// TIA Portal project "Lagerregal_1" (V20)

(* hardware
DEVICE "S7-1500/ET200MP-Station_1"  S7-1500 station
   slot 0: "Profilschiene_0"  Rack  6ES7 590-1***0-0AA0
   slot 1: "PLC_1"  CPU 1513-1 PN  6ES7 513-1AM03-0AB0  V4.0
      slot 3: "CPU-Display_1"  6ES7591-1AA00-0AA0
      slot 32768: "PROFINET-Schnittstelle_1"  X1
         slot 32769: "Port_1"  X1 P1
         slot 32770: "Port_2"  X1 P2
      slot 34817: "Virtual CP interface port_1"  Virtual CP interface port  Virtual CP interface port FW V4.0
   slot 2: "DI 16x24VDC BA_1"  DI 16x24VDC BA  6ES7 521-1BH10-0AA0  V1.1
   slot 3: "DQ 16x24VDC/0.5A ST_1"  DQ 16x24VDC/0.5A ST  6ES7 522-1BH00-0AB0  V2.0
   slot 4: "AI 8xU/I/R/RTD BA_2"  AI 8xU/I/R/RTD BA  6ES7 531-7QF00-0AB0  V1.0
   slot 5: "AI 8xU/I/R/RTD BA_1"  AI 8xU/I/R/RTD BA  6ES7 531-7QF00-0AB0  V1.0
DEVICE "HMI_1"  TP700 Comfort
   slot 0: "HMI_1"  TP700 Comfort  6AV2 124-0GC01-0AX0  17.0.0.0
   slot 1: "HMI_RT_1"  TP700 Comfort  6AV2 124-0GC01-0AX0  17.0.0.0
   slot 5: "HMI_1.IE_CP_1"  PROFINET Interface  17.0.0.0
      slot 1: "PROFINET Schnittstelle_1"  PROFINET Interface
         slot 1: "Port_1"  Port
         slot 2: "Port_2"  Port
   slot 7: "HMI_1.MPI/DP_CP_1"  MPI/DP Interface  17.0.0.0
*)

// ===== PLC "PLC_1"  CPU 1513-1 PN =====

VAR_GLOBAL   // PLC tag table "Variablentabelle aus XML_1"
   "E0.0 Not-Aus (S1)" AT %I0.0 : Bool;
   "E0.1 Anlage ein (S2)" AT %I0.1 : Bool;
   "E0.2 Start (S3)" AT %I0.2 : Bool;
   "E0.3 Sensor_Ein_SS (1B1)" AT %I0.3 : Bool;
   "E0.4 Sensor_Ein_SE (1B2)" AT %I0.4 : Bool;
   "E0.5 Sensor_Ein_MS (2B1)" AT %I0.5 : Bool;
   "E0.6 Sensor_Ein_ME (2B2)" AT %I0.6 : Bool;
   "E0.7 Sensor_Ein_EE (3B1)" AT %I0.7 : Bool;
   "E1.0 Sensor_Aus_S (4B1)" AT %I1.0 : Bool;
   "E1.1 Sensor_Aus_A (5B1)" AT %I1.1 : Bool;
   "E1.2 Kran_Gabel_Endlage (links) (6B1)" AT %I1.2 : Bool;
   "E1.3 Kran_Gabel_Endlage (rechts) (6B2)" AT %I1.3 : Bool;
   "E1.4 Kran_Gabel_Endage (mitte) (6B3)" AT %I1.4 : Bool;
   "E1.5 Kran_Gabel_Endlage (links) (7B1)" AT %I1.5 : Bool;
   "E1.6 Kran_Gabel_Endlage (rechts) (7B2)" AT %I1.6 : Bool;
   "E1.7 Kran_Gabel_Endage (mitte) (7B3)" AT %I1.7 : Bool;
   "A0.2 Start (H3)" AT %Q0.2 : Bool;
   "A0.3 Band_Ein_1 (1M1)" AT %Q0.3 : Bool;
   "A0.5 Band_Ein_2 (2M1)" AT %Q0.5 : Bool;
   "A0.7 Band_Ein_3 (3M1)" AT %Q0.7 : Bool;
   "A1.0 Band_Aus_1 (4M1)" AT %Q1.0 : Bool;
   "A1.1 Band_Aus_2 (5M1)" AT %Q1.1 : Bool;
   "A1.2 Kran_Gabel (links) (6M1)" AT %Q1.2 : Bool;
   "A1.3 Kran_Gabel (rechts) (6M2)" AT %Q1.3 : Bool;
   "A1.5 Kran_Gabel (links) (7M1)" AT %Q1.5 : Bool;
   "A1.6 Kran_Gabel (rechts) (7M2)" AT %Q1.6 : Bool;
   "EW30 Kamera (2B1)" AT %EW30 : Int;
   "EW34 Kran_Ist-X-Pos (6B4)" AT %EW32 : Int;
   "EW38 Kran_Ist-Z-Pos (6B5)" AT %EW34 : Int;
   "EW42 Kran_Ist-X-Pos (7B4)" AT %EW36 : Int;
   "EW46 Kran_Ist-Z-Pos (7B5)" AT %EW38 : Int;
   "AW34 Kran_Soll-X-Pos (6M4)" AT %AW32 : Int;
   "AW38 Kran_Soll-Z-Pos (6M5)" AT %AW34 : Int;
   "AW42 Kran_Soll-X-Pos (7M4)" AT %AW36 : Int;
   "AW46 Kran_Soll-Z-Pos (7M5)" AT %AW38 : Int;
END_VAR

TYPE "typKran_Pos"
   STRUCT
      "X-Ist" : Int;
      "X-Soll" : Int;
      "Z-Ist" : Int;
      "Z-Soll" : Int;
   END_STRUCT;
END_TYPE

TYPE "typLagerplatz"
   STRUCT
      Pos : Struct
         X : Int;
         Z : Int;
      END_STRUCT;
      Flags : Struct
         Belegt : Bool;
         In_Benutzung : Bool;
      END_STRUCT;
   END_STRUCT;
END_TYPE

DATA_BLOCK "IDB_Anlage"   // DB1
{ S7_Optimized_Access := 'TRUE' }
VERSION : 0.1
// stored: InstanceOfName Ein_Anlage
"Ein_Anlage"
BEGIN
END_DATA_BLOCK

DATA_BLOCK "IDB_HMI"   // DB2
{ S7_Optimized_Access := 'TRUE' }
VERSION : 0.1
// stored: InstanceOfName Ein_HMI
"Ein_HMI"
BEGIN
END_DATA_BLOCK

DATA_BLOCK "HMI_Schnittstelle"   // DB100
{ S7_Optimized_Access := 'TRUE' }
VERSION : 0.1
   VAR
      Eingaenge : Struct
         S1 : Bool;
         "1B1" : Bool;
         "1B2" : Bool;
         "2B1" : Bool;
         "2B2" : Bool;
         "3B1" : Bool;
         "4B1" : Bool;
         "5B1" : Bool;
      END_STRUCT;
      Ausgaenge : Struct
         H1 : Bool;
         "1M1" : Bool;
         "2M1" : Bool;
         "3M1" : Bool;
         "4M1" : Bool;
         "5M1" : Bool;
      END_STRUCT;
      Kraene : Struct
         Kran_1 : "typKran_Pos";
         Kran_2 : "typKran_Pos";
      END_STRUCT;
      Lager : Array[0..9] of "typLagerplatz";
      HMI : Struct
         "X-Pos" : Bool;
         "X-Neg" : Bool;
         "Z-Pos" : Bool;
         "Z-Neg" : Bool;
         Inkrement : UInt;
      END_STRUCT;
      Ergebnis : Struct
         "X-Soll" : Int;
         "Z-Soll" : Int;
      END_STRUCT;
   END_VAR
BEGIN
END_DATA_BLOCK

FUNCTION_BLOCK "Ein_Anlage"   // FB1, FBD
{ S7_Optimized_Access := 'TRUE' }
VERSION : 0.1
   VAR
      NTRIG_MDB_1B2 : F_TRIG;
      NTRIG_MDB_2B2 : F_TRIG;
   END_VAR
BEGIN

REGION Network 1: Kran_1 einlesen
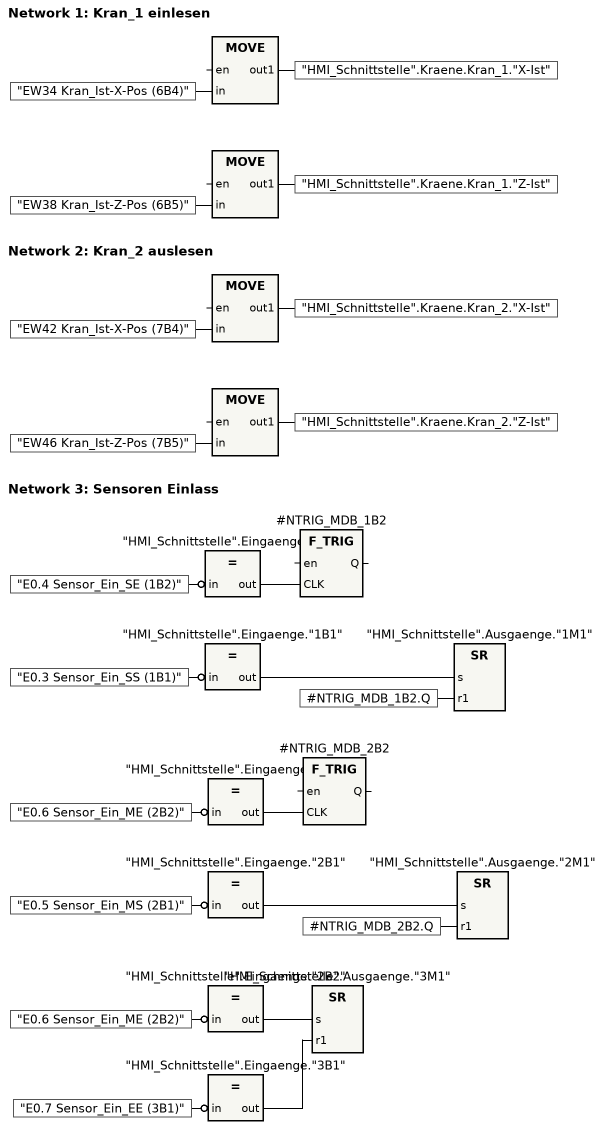
   "HMI_Schnittstelle".Kraene.Kran_1."X-Ist" := "EW34 Kran_Ist-X-Pos (6B4)";
   "HMI_Schnittstelle".Kraene.Kran_1."Z-Ist" := "EW38 Kran_Ist-Z-Pos (6B5)";
END_REGION

REGION Network 2: Kran_2 auslesen
   "HMI_Schnittstelle".Kraene.Kran_2."X-Ist" := "EW42 Kran_Ist-X-Pos (7B4)";
   "HMI_Schnittstelle".Kraene.Kran_2."Z-Ist" := "EW46 Kran_Ist-Z-Pos (7B5)";
END_REGION

REGION Network 3: Sensoren Einlass
   "HMI_Schnittstelle".Eingaenge."1B2" := NOT "E0.4 Sensor_Ein_SE (1B2)";
   #NTRIG_MDB_1B2(CLK := NOT "E0.4 Sensor_Ein_SE (1B2)");   // F_TRIG
   "HMI_Schnittstelle".Eingaenge."1B1" := NOT "E0.3 Sensor_Ein_SS (1B1)";
   IF NOT "E0.3 Sensor_Ein_SS (1B1)" THEN
       "HMI_Schnittstelle".Ausgaenge."1M1" := TRUE;   // SR flip-flop
   END_IF;
   IF #NTRIG_MDB_1B2.Q THEN "HMI_Schnittstelle".Ausgaenge."1M1" := FALSE; END_IF;
   "HMI_Schnittstelle".Eingaenge."2B2" := NOT "E0.6 Sensor_Ein_ME (2B2)";
   #NTRIG_MDB_2B2(CLK := NOT "E0.6 Sensor_Ein_ME (2B2)");   // F_TRIG
   "HMI_Schnittstelle".Eingaenge."2B1" := NOT "E0.5 Sensor_Ein_MS (2B1)";
   IF NOT "E0.5 Sensor_Ein_MS (2B1)" THEN
       "HMI_Schnittstelle".Ausgaenge."2M1" := TRUE;   // SR flip-flop
   END_IF;
   IF #NTRIG_MDB_2B2.Q THEN "HMI_Schnittstelle".Ausgaenge."2M1" := FALSE; END_IF;
   "HMI_Schnittstelle".Eingaenge."2B2" := NOT "E0.6 Sensor_Ein_ME (2B2)";
   "HMI_Schnittstelle".Eingaenge."3B1" := NOT "E0.7 Sensor_Ein_EE (3B1)";
   IF NOT "E0.6 Sensor_Ein_ME (2B2)" THEN
       "HMI_Schnittstelle".Ausgaenge."3M1" := TRUE;   // SR flip-flop
   END_IF;
   IF NOT "E0.7 Sensor_Ein_EE (3B1)" THEN "HMI_Schnittstelle".Ausgaenge."3M1" := FALSE; END_IF;
END_REGION

REGION Network 4 (SCL): Sensoren Auslass
   "HMI_Schnittstelle".Eingaenge."4B1" := NOT "E1.0 Sensor_Aus_S (4B1)";
   "HMI_Schnittstelle".Eingaenge."5B1" := NOT "E1.1 Sensor_Aus_A (5B1)";
END_REGION
END_FUNCTION_BLOCK

FUNCTION_BLOCK "Ein_HMI"   // FB2, FBD
{ S7_Optimized_Access := 'TRUE' }
VERSION : 0.1
   VAR
      "PTRIG_MDB_X-Pos" : R_TRIG;
      "PTRIG_MDB_X-Neg" : R_TRIG;
      "PTRIG_MDB_Z-Pos" : R_TRIG;
      "PTRIG_MDB_Z-Neg" : R_TRIG;
   END_VAR
BEGIN

REGION Network 1
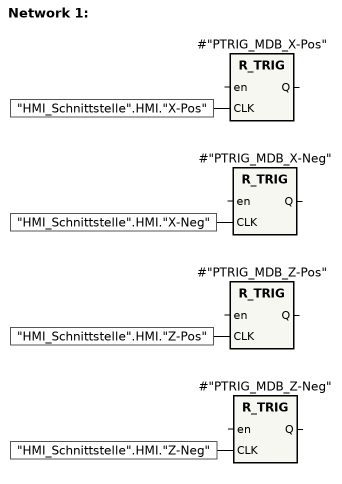
   #"PTRIG_MDB_X-Pos"(CLK := "HMI_Schnittstelle".HMI."X-Pos");   // R_TRIG
   #"PTRIG_MDB_X-Neg"(CLK := "HMI_Schnittstelle".HMI."X-Neg");   // R_TRIG
   #"PTRIG_MDB_Z-Pos"(CLK := "HMI_Schnittstelle".HMI."Z-Pos");   // R_TRIG
   #"PTRIG_MDB_Z-Neg"(CLK := "HMI_Schnittstelle".HMI."Z-Neg");   // R_TRIG
END_REGION
END_FUNCTION_BLOCK

FUNCTION "Aus_Anlage" : Void   // FC1, FBD
{ S7_Optimized_Access := 'TRUE' }
VERSION : 0.1
BEGIN

REGION Network 1: Kran_1 steuern
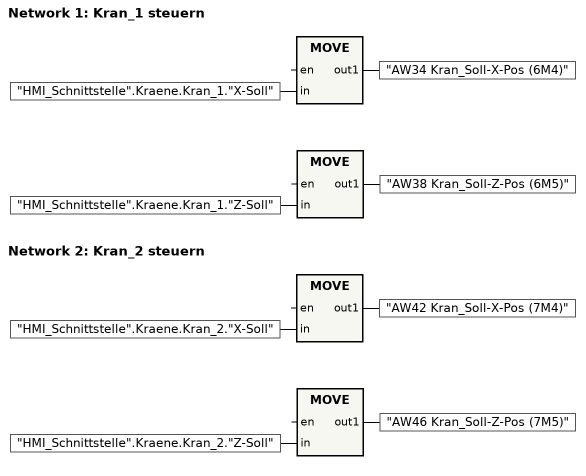
   "AW34 Kran_Soll-X-Pos (6M4)" := "HMI_Schnittstelle".Kraene.Kran_1."X-Soll";
   "AW38 Kran_Soll-Z-Pos (6M5)" := "HMI_Schnittstelle".Kraene.Kran_1."Z-Soll";
END_REGION

REGION Network 2: Kran_2 steuern
   "AW42 Kran_Soll-X-Pos (7M4)" := "HMI_Schnittstelle".Kraene.Kran_2."X-Soll";
   "AW46 Kran_Soll-Z-Pos (7M5)" := "HMI_Schnittstelle".Kraene.Kran_2."Z-Soll";
END_REGION

REGION Network 3 (SCL): Foerderbaender Einlass
   "A0.3 Band_Ein_1 (1M1)" := "HMI_Schnittstelle".Ausgaenge."1M1";
   "A0.5 Band_Ein_2 (2M1)" := "HMI_Schnittstelle".Ausgaenge."2M1";
   "A0.7 Band_Ein_3 (3M1)" := "HMI_Schnittstelle".Ausgaenge."3M1";
END_REGION

REGION Network 4 (SCL): Foerderbaender Auslass
   "A1.0 Band_Aus_1 (4M1)" := "HMI_Schnittstelle".Ausgaenge."4M1";
   "A1.1 Band_Aus_2 (5M1)" := "HMI_Schnittstelle".Ausgaenge."5M1";
END_REGION
END_FUNCTION

FUNCTION "Aus_HMI" : Void   // FC2, FBD
{ S7_Optimized_Access := 'TRUE' }
VERSION : 0.1
BEGIN

REGION Network 2 (SCL): Achsen inkrementieren
   // X-Achse Inkrementieren
   IF "IDB_HMI"."PTRIG_MDB_X-Pos".Q THEN
       "HMI_Schnittstelle".Kraene.Kran_1."X-Soll" += UINT_TO_INT("HMI_Schnittstelle".HMI.Inkrement);
   END_IF;

   IF "IDB_HMI"."PTRIG_MDB_X-Neg".Q THEN
       "HMI_Schnittstelle".Kraene.Kran_1."X-Soll" -= UINT_TO_INT("HMI_Schnittstelle".HMI.Inkrement);
   END_IF;


   // Z-Achse Inkrementieren
   IF "IDB_HMI"."PTRIG_MDB_Z-Pos".Q THEN
       "HMI_Schnittstelle".Kraene.Kran_1."Z-Soll" += UINT_TO_INT("HMI_Schnittstelle".HMI.Inkrement);
   END_IF;

   IF "IDB_HMI"."PTRIG_MDB_Z-Neg".Q THEN
       "HMI_Schnittstelle".Kraene.Kran_1."Z-Soll" -= UINT_TO_INT("HMI_Schnittstelle".HMI.Inkrement);
   END_IF;
END_REGION

REGION Network 3 (SCL): Fachposition berechnen
   //POS_X := ((FachNr - 1) MOD AnzFaecherX) * Facbreite + Off_Null_X;
   //POS_Z := ((FachNr - 1) DIV AnzFaecherX) * Fachoehe + Off_Null_Z;
END_REGION
END_FUNCTION

ORGANIZATION_BLOCK "Main"   // OB1, FBD, ProgramCycle
TITLE = "Main Program Sweep (Cycle)"
{ S7_Optimized_Access := 'TRUE' }
VERSION : 0.1
   VAR_INPUT
      Initial_Call : Bool;   // Initial call of this OB
      Remanence : Bool;   // =True, if remanent data are available
   END_VAR
BEGIN

REGION Network 1: Anlage
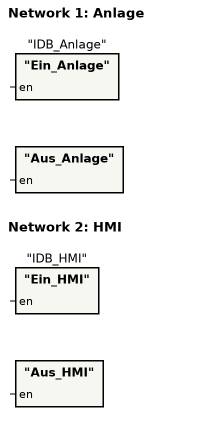
   "IDB_Anlage"();   // "Ein_Anlage"
   "Aus_Anlage"();
END_REGION

REGION Network 2: HMI
   "IDB_HMI"();   // "Ein_HMI"
   "Aus_HMI"();
END_REGION
END_ORGANIZATION_BLOCK

(* ===== HMI "HMI_RT_1" =====
system functions are stored by id; their names below are inferred from use
connection "HMI_Verbindung_1": ETHERNET, S7_1500_OMS

HMI tags "Standard-Variablentabelle"
   "HMI_Schnittstelle_Kraene_Kran_1_Z-Soll" : Int = PLC HMI_Schnittstelle.Kraene.Kran_1.Z-Soll, 1 s
   "HMI_Schnittstelle_Kraene_Kran_1_X-Soll" : Int = PLC HMI_Schnittstelle.Kraene.Kran_1.X-Soll, 1 s
   "HMI_Schnittstelle_Kraene_Kran_1_X-Ist" : Int = PLC HMI_Schnittstelle.Kraene.Kran_1.X-Ist, 1 s
   "HMI_Schnittstelle_Kraene_Kran_1_Z-Ist" : Int = PLC HMI_Schnittstelle.Kraene.Kran_1.Z-Ist, 1 s
   "HMI_Schnittstelle_Lager{0}_Pos_X" : Int = PLC HMI_Schnittstelle.Lager[0].Pos.X, 1 s
   "HMI_Schnittstelle_Lager{0}_Pos_Z" : Int = PLC HMI_Schnittstelle.Lager[0].Pos.Z, 1 s
   "HMI_Schnittstelle_Lager{1}_Pos_X" : Int = PLC HMI_Schnittstelle.Lager[1].Pos.X, 1 s
   "HMI_Schnittstelle_Lager{1}_Pos_Z" : Int = PLC HMI_Schnittstelle.Lager[1].Pos.Z, 1 s
   "HMI_Schnittstelle_Lager{9}_Pos_X" : Int = PLC HMI_Schnittstelle.Lager[9].Pos.X, 1 s
   "HMI_Schnittstelle_Lager{9}_Pos_Z" : Int = PLC HMI_Schnittstelle.Lager[9].Pos.Z, 1 s
   "HMI_Schnittstelle_HMI_X-Neg" : Bool = PLC HMI_Schnittstelle.HMI.X-Neg, 1 s
   "HMI_Schnittstelle_HMI_X-Pos" : Bool = PLC HMI_Schnittstelle.HMI.X-Pos, 1 s
   "HMI_Schnittstelle_HMI_Z-Neg" : Bool = PLC HMI_Schnittstelle.HMI.Z-Neg, 1 s
   "HMI_Schnittstelle_HMI_Z-Pos" : Bool = PLC HMI_Schnittstelle.HMI.Z-Pos, 1 s
   "HMI_Schnittstelle_HMI_Inkrement" : UInt = PLC HMI_Schnittstelle.HMI.Inkrement, 1 s

screen "Lageransicht" 800x420
   Button "Schaltfläche_1" at 100,348 size 64x64; TextOff '9'
   Button "Schaltfläche_2" at 167,348 size 64x64; TextOff '8'
   Button "Schaltfläche_3" at 234,348 size 64x64; TextOff '7'
   Button "Schaltfläche_4" at 10,438 size 96x32; TextOff 'Teachen'
      on Press: ActivateScreen("Teachmodus", 0)
   Button "Schaltfläche_5" at 301,348 size 64x64; TextOff '6'
   Button "Schaltfläche_6" at 368,348 size 64x64; TextOff '5'
   Button "Schaltfläche_7" at 435,348 size 64x64; TextOff '4'
   Button "Schaltfläche_8" at 502,348 size 64x64; TextOff '3'
   Button "Schaltfläche_9" at 569,348 size 64x64; TextOff '2'
   Button "Schaltfläche_10" at 636,348 size 64x64; TextOff '1'
   Button "Schaltfläche_11" at 100,281 size 64x64; TextOff '18'
   Button "Schaltfläche_12" at 167,281 size 64x64; TextOff '17'
   Button "Schaltfläche_13" at 234,281 size 64x64; TextOff '16'
   Button "Schaltfläche_14" at 301,281 size 64x64; TextOff '15'
   Button "Schaltfläche_15" at 368,281 size 64x64; TextOff '14'
   Button "Schaltfläche_16" at 435,281 size 64x64; TextOff '13'
   Button "Schaltfläche_17" at 502,281 size 64x64; TextOff '12'
   Button "Schaltfläche_18" at 569,281 size 64x64; TextOff '11'
   Button "Schaltfläche_19" at 636,281 size 64x64; TextOff '10'
   Button "Schaltfläche_20" at 100,214 size 64x64; TextOff '27'
   Button "Schaltfläche_21" at 167,214 size 64x64; TextOff '26'
   Button "Schaltfläche_22" at 234,214 size 64x64; TextOff '25'
   Button "Schaltfläche_23" at 301,214 size 64x64; TextOff '24'
   Button "Schaltfläche_24" at 368,214 size 64x64; TextOff '23'
   Button "Schaltfläche_25" at 435,214 size 64x64; TextOff '22'
   Button "Schaltfläche_26" at 502,214 size 64x64; TextOff '21'
   Button "Schaltfläche_27" at 569,214 size 64x64; TextOff '20'
   Button "Schaltfläche_28" at 636,214 size 64x64; TextOff '19'
   Button "Schaltfläche_29" at 100,147 size 64x64; TextOff '36'
   Button "Schaltfläche_30" at 167,147 size 64x64; TextOff '35'
   Button "Schaltfläche_31" at 234,147 size 64x64; TextOff '34'
   Button "Schaltfläche_32" at 301,147 size 64x64; TextOff '33'
   Button "Schaltfläche_33" at 368,147 size 64x64; TextOff '32'
   Button "Schaltfläche_34" at 435,147 size 64x64; TextOff '31'
   Button "Schaltfläche_35" at 502,147 size 64x64; TextOff '30'
   Button "Schaltfläche_36" at 569,147 size 64x64; TextOff '29'
   Button "Schaltfläche_37" at 636,147 size 64x64; TextOff '28'
   Button "Schaltfläche_38" at 100,80 size 64x64; TextOff '45'
   Button "Schaltfläche_39" at 167,80 size 64x64; TextOff '44'
   Button "Schaltfläche_40" at 234,80 size 64x64; TextOff '43'
   Button "Schaltfläche_41" at 301,80 size 64x64; TextOff '42'
   Button "Schaltfläche_42" at 368,80 size 64x64; TextOff '41'
   Button "Schaltfläche_43" at 435,80 size 64x64; TextOff '40'
   Button "Schaltfläche_44" at 502,80 size 64x64; TextOff '39'
   Button "Schaltfläche_45" at 569,80 size 64x64; TextOff '38'
   Button "Schaltfläche_46" at 636,80 size 64x64; TextOff '37'
   Button "Schaltfläche_47" at 100,13 size 64x64; TextOff '54'
   Button "Schaltfläche_48" at 167,13 size 64x64; TextOff '53'
   Button "Schaltfläche_49" at 234,13 size 64x64; TextOff '52'
   Button "Schaltfläche_50" at 301,13 size 64x64; TextOff '51'
   Button "Schaltfläche_51" at 368,13 size 64x64; TextOff '50'
   Button "Schaltfläche_52" at 435,13 size 64x64; TextOff '49'
   Button "Schaltfläche_53" at 502,13 size 64x64; TextOff '48'
   Button "Schaltfläche_54" at 569,13 size 64x64; TextOff '47'
   Button "Schaltfläche_55" at 636,13 size 64x64; TextOff '46'

screen "Teachmodus" 800x420, template "Menüleiste"
   Button "Schaltfläche_1" at 694,10 size 96x32; TextOff 'Zurück'
      on Press: function_efd93a16()
   TextField "Textfeld_1" at 308,10 size 184x23; Text 'Kalibrierungsmodus'
   TextField "Textfeld_2" at 670,64 size 119x23; Text 'Lagerplatz 1'
   IOField "EA-Feld_1" at 459,92 size 96x32; FormatPattern 99999
      ProcessValue <- "HMI_Schnittstelle_Lager{0}_Pos_X"
   IOField "EA-Feld_2" at 563,92 size 96x32; FormatPattern 99999
      ProcessValue <- "HMI_Schnittstelle_Lager{0}_Pos_Z"
   TextField "Textfeld_4" at 458,64 size 78x23; Text 'X-Achse'
   TextField "Textfeld_5" at 563,64 size 77x23; Text 'Z-Achse'
   Button "Schaltfläche_2" at 694,92 size 96x32; TextOff 'Bestätigen'
      on Press: SetTag("HMI_Schnittstelle_Lager{0}_Pos_X", "HMI_Schnittstelle_Kraene_Kran_1_X-Ist"); SetTag("HMI_Schnittstelle_Lager{0}_Pos_Z", "HMI_Schnittstelle_Kraene_Kran_1_Z-Ist")
   TextField "Textfeld_3" at 670,139 size 119x23; Text 'Lagerplatz 2'
   IOField "EA-Feld_3" at 459,168 size 96x32; FormatPattern 99999
      ProcessValue <- "HMI_Schnittstelle_Lager{1}_Pos_X"
   IOField "EA-Feld_4" at 563,168 size 96x32; FormatPattern 99999
      ProcessValue <- "HMI_Schnittstelle_Lager{1}_Pos_Z"
   TextField "Textfeld_6" at 458,140 size 78x23; Text 'X-Achse'
   TextField "Textfeld_7" at 563,140 size 77x23; Text 'Z-Achse'
   Button "Schaltfläche_3" at 694,168 size 96x32; TextOff 'Bestätigen'
      on Press: SetTag("HMI_Schnittstelle_Lager{1}_Pos_X", "HMI_Schnittstelle_Kraene_Kran_1_X-Ist"); SetTag("HMI_Schnittstelle_Lager{1}_Pos_Z", "HMI_Schnittstelle_Kraene_Kran_1_Z-Ist")
   TextField "Textfeld_8" at 658,216 size 130x23; Text 'Lagerplatz 10'
   IOField "EA-Feld_5" at 459,244 size 96x32; FormatPattern 99999
      ProcessValue <- "HMI_Schnittstelle_Lager{9}_Pos_X"
   IOField "EA-Feld_6" at 563,244 size 96x32; FormatPattern 99999
      ProcessValue <- "HMI_Schnittstelle_Lager{9}_Pos_Z"
   TextField "Textfeld_9" at 458,216 size 78x23; Text 'X-Achse'
   TextField "Textfeld_10" at 563,216 size 77x23; Text 'Z-Achse'
   Button "Schaltfläche_4" at 694,244 size 96x32; TextOff 'Bestätigen'
      on Press: SetTag("HMI_Schnittstelle_Lager{9}_Pos_X", "HMI_Schnittstelle_Kraene_Kran_1_X-Ist"); SetTag("HMI_Schnittstelle_Lager{9}_Pos_Z", "HMI_Schnittstelle_Kraene_Kran_1_Z-Ist")
   Slider "Schieberegler_2" at 87,300 size 230x50; Caption 'Breite'
      ProcessValue <- "HMI_Schnittstelle_Kraene_Kran_1_X-Soll"
   IOField "EA-Feld_8" at 130,130 size 96x32; FormatPattern 99999
      ProcessValue <- "HMI_Schnittstelle_Kraene_Kran_1_X-Ist"
   IOField "EA-Feld_9" at 130,168 size 96x32; FormatPattern 99999
      ProcessValue <- "HMI_Schnittstelle_Kraene_Kran_1_Z-Ist"
   Slider "Schieberegler_1" at 10,43 size 50x230; Caption 'Höhe'
      ProcessValue <- "HMI_Schnittstelle_Kraene_Kran_1_Z-Soll"
   Button "Schaltfläche_5" at 319,300 size 25x50; TextOff '-'
      on Press: function_b14e0dd5("HMI_Schnittstelle_HMI_X-Neg", 0)
      Appearance <- "HMI_Schnittstelle_HMI_X-Neg"
   Button "Schaltfläche_6" at 60,300 size 25x50; TextOff '+'
      on Press: function_b14e0dd5("HMI_Schnittstelle_HMI_X-Pos", 0)
      Appearance <- "HMI_Schnittstelle_HMI_X-Pos"
   IOField "EA-Feld_7" at 11,301 size 48x48; FormatPattern 999
      ProcessValue <- "HMI_Schnittstelle_HMI_Inkrement"
   Button "Schaltfläche_7" at 10,275 size 50x25; TextOff '-'
      on Press: function_b14e0dd5("HMI_Schnittstelle_HMI_Z-Neg", 0)
      Appearance <- "HMI_Schnittstelle_HMI_Z-Neg"
   Button "Schaltfläche_8" at 10,16 size 50x25; TextOff '+'
      on Press: function_b14e0dd5("HMI_Schnittstelle_HMI_Z-Pos", 0)
      Appearance <- "HMI_Schnittstelle_HMI_Z-Pos"

screen "Detailansicht" 800x420
   Button "Schaltfläche_1" at 10,10 size 96x32; TextOff 'Zurück'
      on Press: function_efd93a16()

Template "Menüleiste" 800x420
   TextField "Vorlage_Textfeld_1" at 358,379 size 104x23; Text 'Menüleiste'
*)